END_REGION

REGION Network 2: EM - Resetting State Complete
   RUNG wire#powerrail
      Contact( "EM02".PackML_Sts.Alarm.sts_Resetting_SC )
      wire#w1
      Contact( "EM02".PackML_Sts.CM01.sts_Resetting_SC )
      wire#w2
      Contact( "EM02".PackML_Sts.CM02.sts_Resetting_SC )
      wire#w3
      Contact( "EM02".PackML_Sts.CM03.sts_Resetting_SC )
      wire#w4
      Contact( "EM02".PackML_Sts.CM04.sts_Resetting_SC )
      wire#w5
      Contact( "EM02".PackML_Sts.CM05.sts_Resetting_SC )
      wire#w6
      Contact( "EM02".PackML_Sts.CM06.sts_Resetting_SC )
      wire#w7
      Contact( "EM02".PackML_Sts.CM07.sts_Resetting_SC )
      wire#w8
      Contact( "EM02".PackML_Sts.CM08.sts_Resetting_SC )
      wire#w9
      Contact( "EM02".PackML_Sts.CM09.sts_Resetting_SC )
      wire#w10
      Contact( "EM02".PackML_Sts.CM10.sts_Resetting_SC )
      wire#w11
      Coil( "EM02".PackML_Sts.Unit.sts_Resetting_SC )
   END_RUNG
   RUNG wire#powerrail
      I_Contact( "EM02".PackML_Sts.Alarm.moduleActive )
   END_RUNG wire#w1
   RUNG wire#w1
      I_Contact( "EM02".PackML_Sts.CM01.moduleActive )
   END_RUNG wire#w2
   RUNG wire#w2
      I_Contact( "EM02".PackML_Sts.CM02.moduleActive )
   END_RUNG wire#w3
   RUNG wire#w3
      I_Contact( "EM02".PackML_Sts.CM03.moduleActive )
   END_RUNG wire#w4
   RUNG wire#w4
      I_Contact( "EM02".PackML_Sts.CM04.moduleActive )
   END_RUNG wire#w5
   RUNG wire#w5
      I_Contact( "EM02".PackML_Sts.CM05.moduleActive )
   END_RUNG wire#w6
   RUNG wire#w6
      I_Contact( "EM02".PackML_Sts.CM06.moduleActive )
   END_RUNG wire#w7
   RUNG wire#w7
      I_Contact( "EM02".PackML_Sts.CM07.moduleActive )
   END_RUNG wire#w8
   RUNG wire#w8
      I_Contact( "EM02".PackML_Sts.CM08.moduleActive )
   END_RUNG wire#w9
   RUNG wire#w9
      I_Contact( "EM02".PackML_Sts.CM09.moduleActive )
   END_RUNG wire#w10
   RUNG wire#w10
      I_Contact( "EM02".PackML_Sts.CM10.moduleActive )
   END_RUNG wire#w11
   // the same network as SCL:
   "EM02".PackML_Sts.Unit.sts_Resetting_SC := ("EM02".PackML_Sts.Alarm.sts_Resetting_SC OR NOT "EM02".PackML_Sts.Alarm.moduleActive) AND ("EM02".PackML_Sts.CM01.sts_Resetting_SC OR NOT "EM02".PackML_Sts.CM01.moduleActive) AND ("EM02".PackML_Sts.CM02.sts_Resetting_SC OR NOT "EM02".PackML_Sts.CM02.moduleActive) AND ("EM02".PackML_Sts.CM03.sts_Resetting_SC OR NOT "EM02".PackML_Sts.CM03.moduleActive) AND ("EM02".PackML_Sts.CM04.sts_Resetting_SC OR NOT "EM02".PackML_Sts.CM04.moduleActive) AND ("EM02".PackML_Sts.CM05.sts_Resetting_SC OR NOT "EM02".PackML_Sts.CM05.moduleActive) AND ("EM02".PackML_Sts.CM06.sts_Resetting_SC OR NOT "EM02".PackML_Sts.CM06.moduleActive) AND ("EM02".PackML_Sts.CM07.sts_Resetting_SC OR NOT "EM02".PackML_Sts.CM07.moduleActive) AND ("EM02".PackML_Sts.CM08.sts_Resetting_SC OR NOT "EM02".PackML_Sts.CM08.moduleActive) AND ("EM02".PackML_Sts.CM09.sts_Resetting_SC OR NOT "EM02".PackML_Sts.CM09.moduleActive) AND ("EM02".PackML_Sts.CM10.sts_Resetting_SC OR NOT "EM02".PackML_Sts.CM10.moduleActive);
END_REGION

REGION Network 3: EM - Start Command
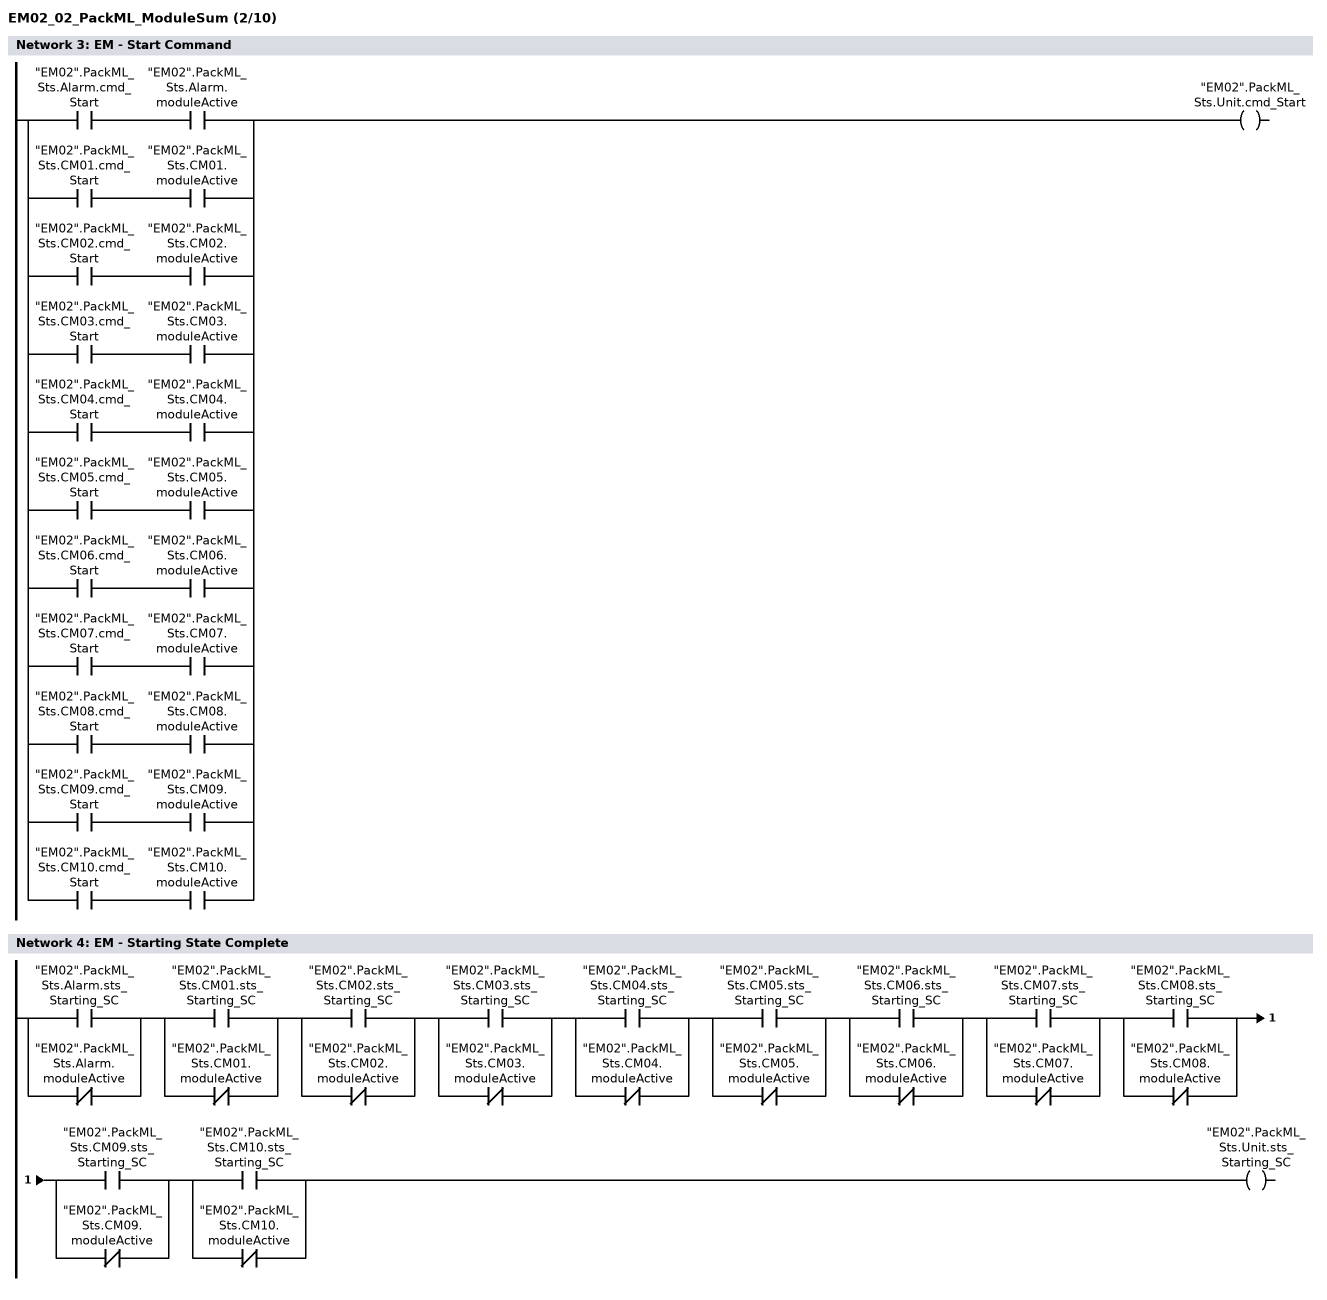
   RUNG wire#powerrail
      Contact( "EM02".PackML_Sts.Alarm.cmd_Start )
      Contact( "EM02".PackML_Sts.Alarm.moduleActive )
      wire#w1
      Coil( "EM02".PackML_Sts.Unit.cmd_Start )
   END_RUNG
   RUNG wire#powerrail
      Contact( "EM02".PackML_Sts.CM01.cmd_Start )
      Contact( "EM02".PackML_Sts.CM01.moduleActive )
   END_RUNG wire#w1
   RUNG wire#powerrail
      Contact( "EM02".PackML_Sts.CM02.cmd_Start )
      Contact( "EM02".PackML_Sts.CM02.moduleActive )
   END_RUNG wire#w1
   RUNG wire#powerrail
      Contact( "EM02".PackML_Sts.CM03.cmd_Start )
      Contact( "EM02".PackML_Sts.CM03.moduleActive )
   END_RUNG wire#w1
   RUNG wire#powerrail
      Contact( "EM02".PackML_Sts.CM04.cmd_Start )
      Contact( "EM02".PackML_Sts.CM04.moduleActive )
   END_RUNG wire#w1
   RUNG wire#powerrail
      Contact( "EM02".PackML_Sts.CM05.cmd_Start )
      Contact( "EM02".PackML_Sts.CM05.moduleActive )
   END_RUNG wire#w1
   RUNG wire#powerrail
      Contact( "EM02".PackML_Sts.CM06.cmd_Start )
      Contact( "EM02".PackML_Sts.CM06.moduleActive )
   END_RUNG wire#w1
   RUNG wire#powerrail
      Contact( "EM02".PackML_Sts.CM07.cmd_Start )
      Contact( "EM02".PackML_Sts.CM07.moduleActive )
   END_RUNG wire#w1
   RUNG wire#powerrail
      Contact( "EM02".PackML_Sts.CM08.cmd_Start )
      Contact( "EM02".PackML_Sts.CM08.moduleActive )
   END_RUNG wire#w1
   RUNG wire#powerrail
      Contact( "EM02".PackML_Sts.CM09.cmd_Start )
      Contact( "EM02".PackML_Sts.CM09.moduleActive )
   END_RUNG wire#w1
   RUNG wire#powerrail
      Contact( "EM02".PackML_Sts.CM10.cmd_Start )
      Contact( "EM02".PackML_Sts.CM10.moduleActive )
   END_RUNG wire#w1
   // the same network as SCL:
   "EM02".PackML_Sts.Unit.cmd_Start := ("EM02".PackML_Sts.Alarm.cmd_Start AND "EM02".PackML_Sts.Alarm.moduleActive) OR ("EM02".PackML_Sts.CM01.cmd_Start AND "EM02".PackML_Sts.CM01.moduleActive) OR ("EM02".PackML_Sts.CM02.cmd_Start AND "EM02".PackML_Sts.CM02.moduleActive) OR ("EM02".PackML_Sts.CM03.cmd_Start AND "EM02".PackML_Sts.CM03.moduleActive) OR ("EM02".PackML_Sts.CM04.cmd_Start AND "EM02".PackML_Sts.CM04.moduleActive) OR ("EM02".PackML_Sts.CM05.cmd_Start AND "EM02".PackML_Sts.CM05.moduleActive) OR ("EM02".PackML_Sts.CM06.cmd_Start AND "EM02".PackML_Sts.CM06.moduleActive) OR ("EM02".PackML_Sts.CM07.cmd_Start AND "EM02".PackML_Sts.CM07.moduleActive) OR ("EM02".PackML_Sts.CM08.cmd_Start AND "EM02".PackML_Sts.CM08.moduleActive) OR ("EM02".PackML_Sts.CM09.cmd_Start AND "EM02".PackML_Sts.CM09.moduleActive) OR ("EM02".PackML_Sts.CM10.cmd_Start AND "EM02".PackML_Sts.CM10.moduleActive);
END_REGION

REGION Network 4: EM - Starting State Complete
   RUNG wire#powerrail
      Contact( "EM02".PackML_Sts.Alarm.sts_Starting_SC )
      wire#w1
      Contact( "EM02".PackML_Sts.CM01.sts_Starting_SC )
      wire#w2
      Contact( "EM02".PackML_Sts.CM02.sts_Starting_SC )
      wire#w3
      Contact( "EM02".PackML_Sts.CM03.sts_Starting_SC )
      wire#w4
      Contact( "EM02".PackML_Sts.CM04.sts_Starting_SC )
      wire#w5
      Contact( "EM02".PackML_Sts.CM05.sts_Starting_SC )
      wire#w6
      Contact( "EM02".PackML_Sts.CM06.sts_Starting_SC )
      wire#w7
      Contact( "EM02".PackML_Sts.CM07.sts_Starting_SC )
      wire#w8
      Contact( "EM02".PackML_Sts.CM08.sts_Starting_SC )
      wire#w9
      Contact( "EM02".PackML_Sts.CM09.sts_Starting_SC )
      wire#w10
      Contact( "EM02".PackML_Sts.CM10.sts_Starting_SC )
      wire#w11
      Coil( "EM02".PackML_Sts.Unit.sts_Starting_SC )
   END_RUNG
   RUNG wire#powerrail
      I_Contact( "EM02".PackML_Sts.Alarm.moduleActive )
   END_RUNG wire#w1
   RUNG wire#w1
      I_Contact( "EM02".PackML_Sts.CM01.moduleActive )
   END_RUNG wire#w2
   RUNG wire#w2
      I_Contact( "EM02".PackML_Sts.CM02.moduleActive )
   END_RUNG wire#w3
   RUNG wire#w3
      I_Contact( "EM02".PackML_Sts.CM03.moduleActive )
   END_RUNG wire#w4
   RUNG wire#w4
      I_Contact( "EM02".PackML_Sts.CM04.moduleActive )
   END_RUNG wire#w5
   RUNG wire#w5
      I_Contact( "EM02".PackML_Sts.CM05.moduleActive )
   END_RUNG wire#w6
   RUNG wire#w6
      I_Contact( "EM02".PackML_Sts.CM06.moduleActive )
   END_RUNG wire#w7
   RUNG wire#w7
      I_Contact( "EM02".PackML_Sts.CM07.moduleActive )
   END_RUNG wire#w8
   RUNG wire#w8
      I_Contact( "EM02".PackML_Sts.CM08.moduleActive )
   END_RUNG wire#w9
   RUNG wire#w9
      I_Contact( "EM02".PackML_Sts.CM09.moduleActive )
   END_RUNG wire#w10
   RUNG wire#w10
      I_Contact( "EM02".PackML_Sts.CM10.moduleActive )
   END_RUNG wire#w11
   // the same network as SCL:
   "EM02".PackML_Sts.Unit.sts_Starting_SC := ("EM02".PackML_Sts.Alarm.sts_Starting_SC OR NOT "EM02".PackML_Sts.Alarm.moduleActive) AND ("EM02".PackML_Sts.CM01.sts_Starting_SC OR NOT "EM02".PackML_Sts.CM01.moduleActive) AND ("EM02".PackML_Sts.CM02.sts_Starting_SC OR NOT "EM02".PackML_Sts.CM02.moduleActive) AND ("EM02".PackML_Sts.CM03.sts_Starting_SC OR NOT "EM02".PackML_Sts.CM03.moduleActive) AND ("EM02".PackML_Sts.CM04.sts_Starting_SC OR NOT "EM02".PackML_Sts.CM04.moduleActive) AND ("EM02".PackML_Sts.CM05.sts_Starting_SC OR NOT "EM02".PackML_Sts.CM05.moduleActive) AND ("EM02".PackML_Sts.CM06.sts_Starting_SC OR NOT "EM02".PackML_Sts.CM06.moduleActive) AND ("EM02".PackML_Sts.CM07.sts_Starting_SC OR NOT "EM02".PackML_Sts.CM07.moduleActive) AND ("EM02".PackML_Sts.CM08.sts_Starting_SC OR NOT "EM02".PackML_Sts.CM08.moduleActive) AND ("EM02".PackML_Sts.CM09.sts_Starting_SC OR NOT "EM02".PackML_Sts.CM09.moduleActive) AND ("EM02".PackML_Sts.CM10.sts_Starting_SC OR NOT "EM02".PackML_Sts.CM10.moduleActive);
END_REGION

REGION Network 5: EM - Stop Command
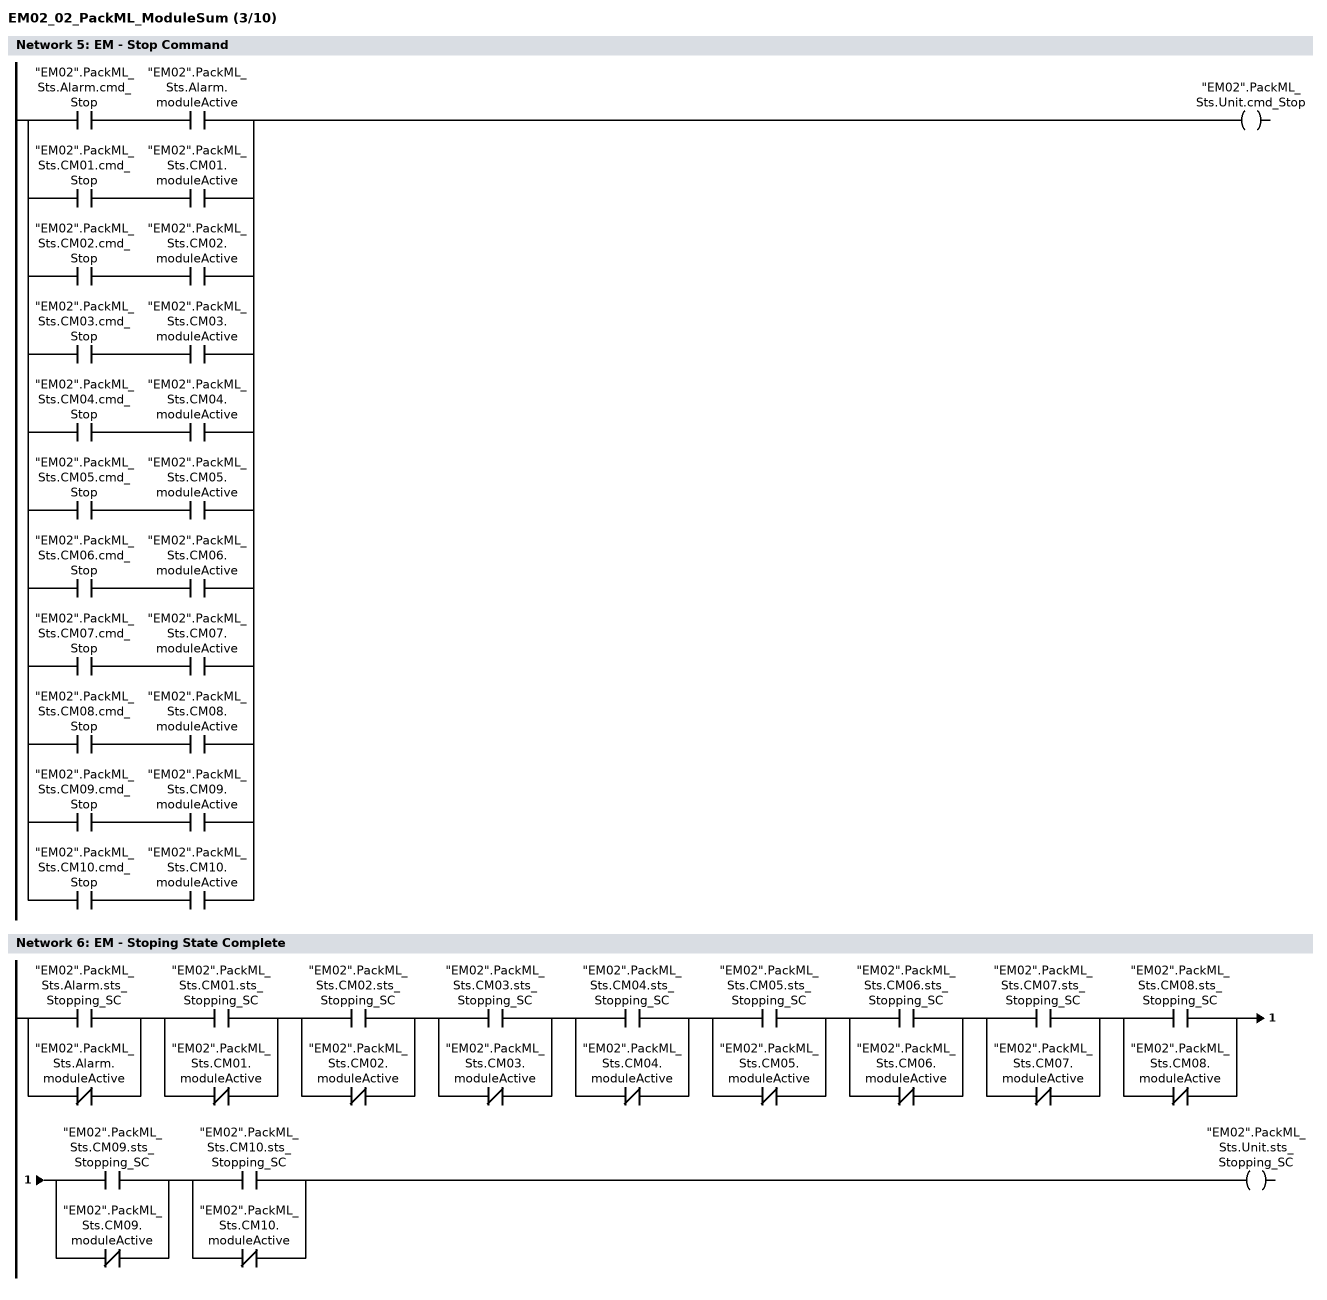
   RUNG wire#powerrail
      Contact( "EM02".PackML_Sts.Alarm.cmd_Stop )
      Contact( "EM02".PackML_Sts.Alarm.moduleActive )
      wire#w1
      Coil( "EM02".PackML_Sts.Unit.cmd_Stop )
   END_RUNG
   RUNG wire#powerrail
      Contact( "EM02".PackML_Sts.CM01.cmd_Stop )
      Contact( "EM02".PackML_Sts.CM01.moduleActive )
   END_RUNG wire#w1
   RUNG wire#powerrail
      Contact( "EM02".PackML_Sts.CM02.cmd_Stop )
      Contact( "EM02".PackML_Sts.CM02.moduleActive )
   END_RUNG wire#w1
   RUNG wire#powerrail
      Contact( "EM02".PackML_Sts.CM03.cmd_Stop )
      Contact( "EM02".PackML_Sts.CM03.moduleActive )
   END_RUNG wire#w1
   RUNG wire#powerrail
      Contact( "EM02".PackML_Sts.CM04.cmd_Stop )
      Contact( "EM02".PackML_Sts.CM04.moduleActive )
   END_RUNG wire#w1
   RUNG wire#powerrail
      Contact( "EM02".PackML_Sts.CM05.cmd_Stop )
      Contact( "EM02".PackML_Sts.CM05.moduleActive )
   END_RUNG wire#w1
   RUNG wire#powerrail
      Contact( "EM02".PackML_Sts.CM06.cmd_Stop )
      Contact( "EM02".PackML_Sts.CM06.moduleActive )
   END_RUNG wire#w1
   RUNG wire#powerrail
      Contact( "EM02".PackML_Sts.CM07.cmd_Stop )
      Contact( "EM02".PackML_Sts.CM07.moduleActive )
   END_RUNG wire#w1
   RUNG wire#powerrail
      Contact( "EM02".PackML_Sts.CM08.cmd_Stop )
      Contact( "EM02".PackML_Sts.CM08.moduleActive )
   END_RUNG wire#w1
   RUNG wire#powerrail
      Contact( "EM02".PackML_Sts.CM09.cmd_Stop )
      Contact( "EM02".PackML_Sts.CM09.moduleActive )
   END_RUNG wire#w1
   RUNG wire#powerrail
      Contact( "EM02".PackML_Sts.CM10.cmd_Stop )
      Contact( "EM02".PackML_Sts.CM10.moduleActive )
   END_RUNG wire#w1
   // the same network as SCL:
   "EM02".PackML_Sts.Unit.cmd_Stop := ("EM02".PackML_Sts.Alarm.cmd_Stop AND "EM02".PackML_Sts.Alarm.moduleActive) OR ("EM02".PackML_Sts.CM01.cmd_Stop AND "EM02".PackML_Sts.CM01.moduleActive) OR ("EM02".PackML_Sts.CM02.cmd_Stop AND "EM02".PackML_Sts.CM02.moduleActive) OR ("EM02".PackML_Sts.CM03.cmd_Stop AND "EM02".PackML_Sts.CM03.moduleActive) OR ("EM02".PackML_Sts.CM04.cmd_Stop AND "EM02".PackML_Sts.CM04.moduleActive) OR ("EM02".PackML_Sts.CM05.cmd_Stop AND "EM02".PackML_Sts.CM05.moduleActive) OR ("EM02".PackML_Sts.CM06.cmd_Stop AND "EM02".PackML_Sts.CM06.moduleActive) OR ("EM02".PackML_Sts.CM07.cmd_Stop AND "EM02".PackML_Sts.CM07.moduleActive) OR ("EM02".PackML_Sts.CM08.cmd_Stop AND "EM02".PackML_Sts.CM08.moduleActive) OR ("EM02".PackML_Sts.CM09.cmd_Stop AND "EM02".PackML_Sts.CM09.moduleActive) OR ("EM02".PackML_Sts.CM10.cmd_Stop AND "EM02".PackML_Sts.CM10.moduleActive);
END_REGION

REGION Network 6: EM - Stoping State Complete
   RUNG wire#powerrail
      Contact( "EM02".PackML_Sts.Alarm.sts_Stopping_SC )
      wire#w1
      Contact( "EM02".PackML_Sts.CM01.sts_Stopping_SC )
      wire#w2
      Contact( "EM02".PackML_Sts.CM02.sts_Stopping_SC )
      wire#w3
      Contact( "EM02".PackML_Sts.CM03.sts_Stopping_SC )
      wire#w4
      Contact( "EM02".PackML_Sts.CM04.sts_Stopping_SC )
      wire#w5
      Contact( "EM02".PackML_Sts.CM05.sts_Stopping_SC )
      wire#w6
      Contact( "EM02".PackML_Sts.CM06.sts_Stopping_SC )
      wire#w7
      Contact( "EM02".PackML_Sts.CM07.sts_Stopping_SC )
      wire#w8
      Contact( "EM02".PackML_Sts.CM08.sts_Stopping_SC )
      wire#w9
      Contact( "EM02".PackML_Sts.CM09.sts_Stopping_SC )
      wire#w10
      Contact( "EM02".PackML_Sts.CM10.sts_Stopping_SC )
      wire#w11
      Coil( "EM02".PackML_Sts.Unit.sts_Stopping_SC )
   END_RUNG
   RUNG wire#powerrail
      I_Contact( "EM02".PackML_Sts.Alarm.moduleActive )
   END_RUNG wire#w1
   RUNG wire#w1
      I_Contact( "EM02".PackML_Sts.CM01.moduleActive )
   END_RUNG wire#w2
   RUNG wire#w2
      I_Contact( "EM02".PackML_Sts.CM02.moduleActive )
   END_RUNG wire#w3
   RUNG wire#w3
      I_Contact( "EM02".PackML_Sts.CM03.moduleActive )
   END_RUNG wire#w4
   RUNG wire#w4
      I_Contact( "EM02".PackML_Sts.CM04.moduleActive )
   END_RUNG wire#w5
   RUNG wire#w5
      I_Contact( "EM02".PackML_Sts.CM05.moduleActive )
   END_RUNG wire#w6
   RUNG wire#w6
      I_Contact( "EM02".PackML_Sts.CM06.moduleActive )
   END_RUNG wire#w7
   RUNG wire#w7
      I_Contact( "EM02".PackML_Sts.CM07.moduleActive )
   END_RUNG wire#w8
   RUNG wire#w8
      I_Contact( "EM02".PackML_Sts.CM08.moduleActive )
   END_RUNG wire#w9
   RUNG wire#w9
      I_Contact( "EM02".PackML_Sts.CM09.moduleActive )
   END_RUNG wire#w10
   RUNG wire#w10
      I_Contact( "EM02".PackML_Sts.CM10.moduleActive )
   END_RUNG wire#w11
   // the same network as SCL:
   "EM02".PackML_Sts.Unit.sts_Stopping_SC := ("EM02".PackML_Sts.Alarm.sts_Stopping_SC OR NOT "EM02".PackML_Sts.Alarm.moduleActive) AND ("EM02".PackML_Sts.CM01.sts_Stopping_SC OR NOT "EM02".PackML_Sts.CM01.moduleActive) AND ("EM02".PackML_Sts.CM02.sts_Stopping_SC OR NOT "EM02".PackML_Sts.CM02.moduleActive) AND ("EM02".PackML_Sts.CM03.sts_Stopping_SC OR NOT "EM02".PackML_Sts.CM03.moduleActive) AND ("EM02".PackML_Sts.CM04.sts_Stopping_SC OR NOT "EM02".PackML_Sts.CM04.moduleActive) AND ("EM02".PackML_Sts.CM05.sts_Stopping_SC OR NOT "EM02".PackML_Sts.CM05.moduleActive) AND ("EM02".PackML_Sts.CM06.sts_Stopping_SC OR NOT "EM02".PackML_Sts.CM06.moduleActive) AND ("EM02".PackML_Sts.CM07.sts_Stopping_SC OR NOT "EM02".PackML_Sts.CM07.moduleActive) AND ("EM02".PackML_Sts.CM08.sts_Stopping_SC OR NOT "EM02".PackML_Sts.CM08.moduleActive) AND ("EM02".PackML_Sts.CM09.sts_Stopping_SC OR NOT "EM02".PackML_Sts.CM09.moduleActive) AND ("EM02".PackML_Sts.CM10.sts_Stopping_SC OR NOT "EM02".PackML_Sts.CM10.moduleActive);
END_REGION

REGION Network 7: EM - Hold Command
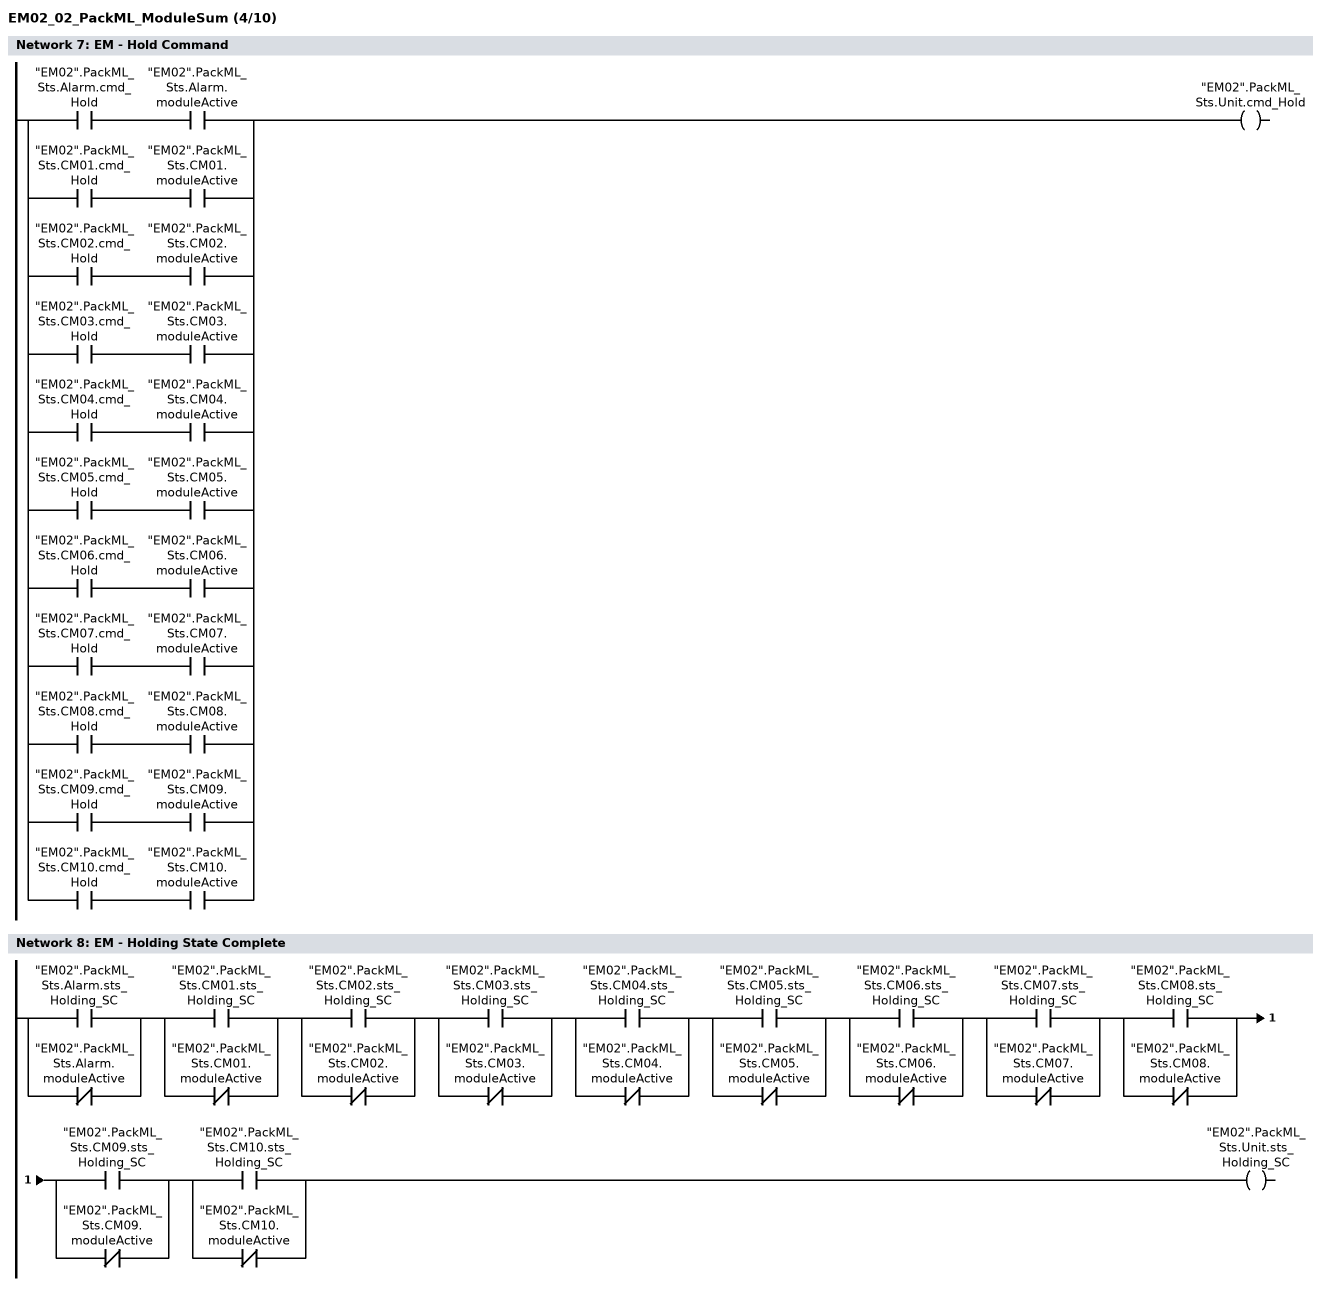
   RUNG wire#powerrail
      Contact( "EM02".PackML_Sts.Alarm.cmd_Hold )
      Contact( "EM02".PackML_Sts.Alarm.moduleActive )
      wire#w1
      Coil( "EM02".PackML_Sts.Unit.cmd_Hold )
   END_RUNG
   RUNG wire#powerrail
      Contact( "EM02".PackML_Sts.CM01.cmd_Hold )
      Contact( "EM02".PackML_Sts.CM01.moduleActive )
   END_RUNG wire#w1
   RUNG wire#powerrail
      Contact( "EM02".PackML_Sts.CM02.cmd_Hold )
      Contact( "EM02".PackML_Sts.CM02.moduleActive )
   END_RUNG wire#w1
   RUNG wire#powerrail
      Contact( "EM02".PackML_Sts.CM03.cmd_Hold )
      Contact( "EM02".PackML_Sts.CM03.moduleActive )
   END_RUNG wire#w1
   RUNG wire#powerrail
      Contact( "EM02".PackML_Sts.CM04.cmd_Hold )
      Contact( "EM02".PackML_Sts.CM04.moduleActive )
   END_RUNG wire#w1
   RUNG wire#powerrail
      Contact( "EM02".PackML_Sts.CM05.cmd_Hold )
      Contact( "EM02".PackML_Sts.CM05.moduleActive )
   END_RUNG wire#w1
   RUNG wire#powerrail
      Contact( "EM02".PackML_Sts.CM06.cmd_Hold )
      Contact( "EM02".PackML_Sts.CM06.moduleActive )
   END_RUNG wire#w1
   RUNG wire#powerrail
      Contact( "EM02".PackML_Sts.CM07.cmd_Hold )
      Contact( "EM02".PackML_Sts.CM07.moduleActive )
   END_RUNG wire#w1
   RUNG wire#powerrail
      Contact( "EM02".PackML_Sts.CM08.cmd_Hold )
      Contact( "EM02".PackML_Sts.CM08.moduleActive )
   END_RUNG wire#w1
   RUNG wire#powerrail
      Contact( "EM02".PackML_Sts.CM09.cmd_Hold )
      Contact( "EM02".PackML_Sts.CM09.moduleActive )
   END_RUNG wire#w1
   RUNG wire#powerrail
      Contact( "EM02".PackML_Sts.CM10.cmd_Hold )
      Contact( "EM02".PackML_Sts.CM10.moduleActive )
   END_RUNG wire#w1
   // the same network as SCL:
   "EM02".PackML_Sts.Unit.cmd_Hold := ("EM02".PackML_Sts.Alarm.cmd_Hold AND "EM02".PackML_Sts.Alarm.moduleActive) OR ("EM02".PackML_Sts.CM01.cmd_Hold AND "EM02".PackML_Sts.CM01.moduleActive) OR ("EM02".PackML_Sts.CM02.cmd_Hold AND "EM02".PackML_Sts.CM02.moduleActive) OR ("EM02".PackML_Sts.CM03.cmd_Hold AND "EM02".PackML_Sts.CM03.moduleActive) OR ("EM02".PackML_Sts.CM04.cmd_Hold AND "EM02".PackML_Sts.CM04.moduleActive) OR ("EM02".PackML_Sts.CM05.cmd_Hold AND "EM02".PackML_Sts.CM05.moduleActive) OR ("EM02".PackML_Sts.CM06.cmd_Hold AND "EM02".PackML_Sts.CM06.moduleActive) OR ("EM02".PackML_Sts.CM07.cmd_Hold AND "EM02".PackML_Sts.CM07.moduleActive) OR ("EM02".PackML_Sts.CM08.cmd_Hold AND "EM02".PackML_Sts.CM08.moduleActive) OR ("EM02".PackML_Sts.CM09.cmd_Hold AND "EM02".PackML_Sts.CM09.moduleActive) OR ("EM02".PackML_Sts.CM10.cmd_Hold AND "EM02".PackML_Sts.CM10.moduleActive);
END_REGION

REGION Network 8: EM - Holding State Complete
   RUNG wire#powerrail
      Contact( "EM02".PackML_Sts.Alarm.sts_Holding_SC )
      wire#w1
      Contact( "EM02".PackML_Sts.CM01.sts_Holding_SC )
      wire#w2
      Contact( "EM02".PackML_Sts.CM02.sts_Holding_SC )
      wire#w3
      Contact( "EM02".PackML_Sts.CM03.sts_Holding_SC )
      wire#w4
      Contact( "EM02".PackML_Sts.CM04.sts_Holding_SC )
      wire#w5
      Contact( "EM02".PackML_Sts.CM05.sts_Holding_SC )
      wire#w6
      Contact( "EM02".PackML_Sts.CM06.sts_Holding_SC )
      wire#w7
      Contact( "EM02".PackML_Sts.CM07.sts_Holding_SC )
      wire#w8
      Contact( "EM02".PackML_Sts.CM08.sts_Holding_SC )
      wire#w9
      Contact( "EM02".PackML_Sts.CM09.sts_Holding_SC )
      wire#w10
      Contact( "EM02".PackML_Sts.CM10.sts_Holding_SC )
      wire#w11
      Coil( "EM02".PackML_Sts.Unit.sts_Holding_SC )
   END_RUNG
   RUNG wire#powerrail
      I_Contact( "EM02".PackML_Sts.Alarm.moduleActive )
   END_RUNG wire#w1
   RUNG wire#w1
      I_Contact( "EM02".PackML_Sts.CM01.moduleActive )
   END_RUNG wire#w2
   RUNG wire#w2
      I_Contact( "EM02".PackML_Sts.CM02.moduleActive )
   END_RUNG wire#w3
   RUNG wire#w3
      I_Contact( "EM02".PackML_Sts.CM03.moduleActive )
   END_RUNG wire#w4
   RUNG wire#w4
      I_Contact( "EM02".PackML_Sts.CM04.moduleActive )
   END_RUNG wire#w5
   RUNG wire#w5
      I_Contact( "EM02".PackML_Sts.CM05.moduleActive )
   END_RUNG wire#w6
   RUNG wire#w6
      I_Contact( "EM02".PackML_Sts.CM06.moduleActive )
   END_RUNG wire#w7
   RUNG wire#w7
      I_Contact( "EM02".PackML_Sts.CM07.moduleActive )
   END_RUNG wire#w8
   RUNG wire#w8
      I_Contact( "EM02".PackML_Sts.CM08.moduleActive )
   END_RUNG wire#w9
   RUNG wire#w9
      I_Contact( "EM02".PackML_Sts.CM09.moduleActive )
   END_RUNG wire#w10
   RUNG wire#w10
      I_Contact( "EM02".PackML_Sts.CM10.moduleActive )
   END_RUNG wire#w11
   // the same network as SCL:
   "EM02".PackML_Sts.Unit.sts_Holding_SC := ("EM02".PackML_Sts.Alarm.sts_Holding_SC OR NOT "EM02".PackML_Sts.Alarm.moduleActive) AND ("EM02".PackML_Sts.CM01.sts_Holding_SC OR NOT "EM02".PackML_Sts.CM01.moduleActive) AND ("EM02".PackML_Sts.CM02.sts_Holding_SC OR NOT "EM02".PackML_Sts.CM02.moduleActive) AND ("EM02".PackML_Sts.CM03.sts_Holding_SC OR NOT "EM02".PackML_Sts.CM03.moduleActive) AND ("EM02".PackML_Sts.CM04.sts_Holding_SC OR NOT "EM02".PackML_Sts.CM04.moduleActive) AND ("EM02".PackML_Sts.CM05.sts_Holding_SC OR NOT "EM02".PackML_Sts.CM05.moduleActive) AND ("EM02".PackML_Sts.CM06.sts_Holding_SC OR NOT "EM02".PackML_Sts.CM06.moduleActive) AND ("EM02".PackML_Sts.CM07.sts_Holding_SC OR NOT "EM02".PackML_Sts.CM07.moduleActive) AND ("EM02".PackML_Sts.CM08.sts_Holding_SC OR NOT "EM02".PackML_Sts.CM08.moduleActive) AND ("EM02".PackML_Sts.CM09.sts_Holding_SC OR NOT "EM02".PackML_Sts.CM09.moduleActive) AND ("EM02".PackML_Sts.CM10.sts_Holding_SC OR NOT "EM02".PackML_Sts.CM10.moduleActive);
END_REGION

REGION Network 9: EM - UnHold Command
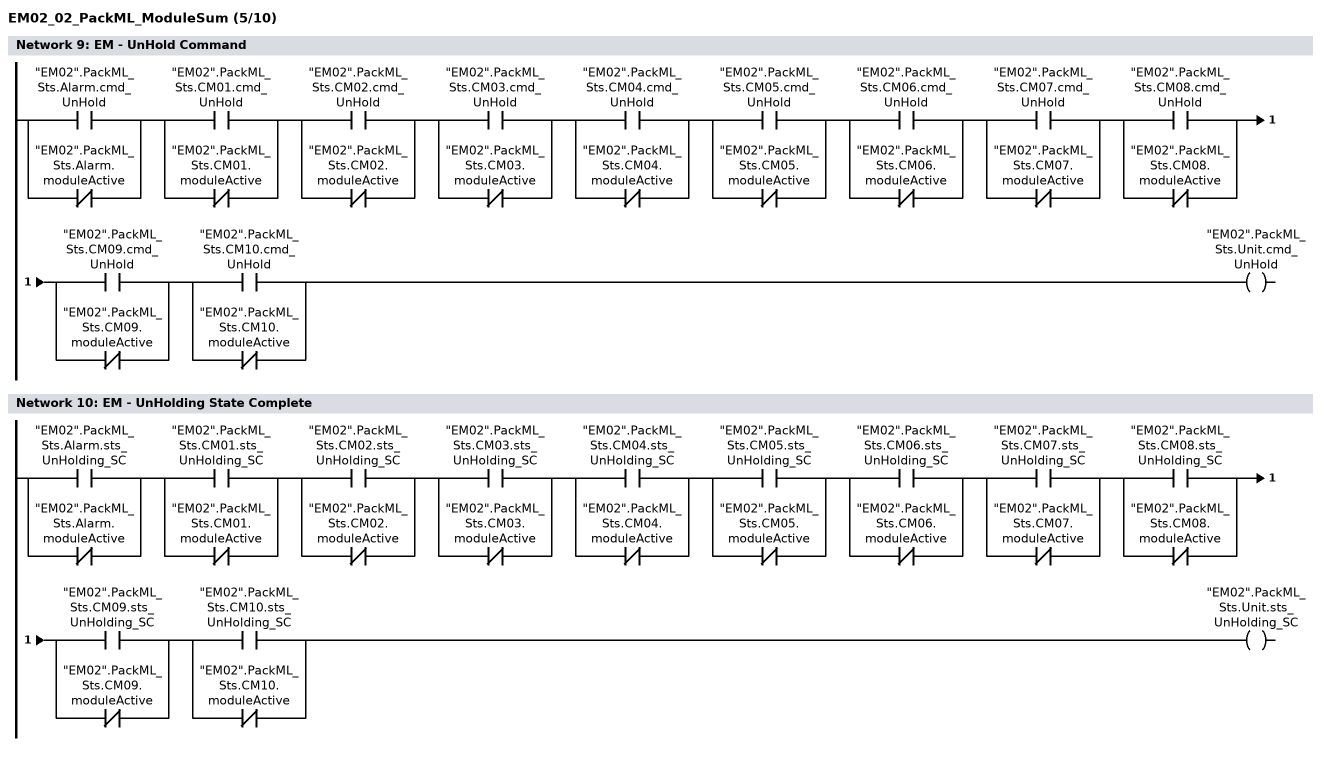
   RUNG wire#powerrail
      Contact( "EM02".PackML_Sts.Alarm.cmd_UnHold )
      wire#w1
      Contact( "EM02".PackML_Sts.CM01.cmd_UnHold )
      wire#w2
      Contact( "EM02".PackML_Sts.CM02.cmd_UnHold )
      wire#w3
      Contact( "EM02".PackML_Sts.CM03.cmd_UnHold )
      wire#w4
      Contact( "EM02".PackML_Sts.CM04.cmd_UnHold )
      wire#w5
      Contact( "EM02".PackML_Sts.CM05.cmd_UnHold )
      wire#w6
      Contact( "EM02".PackML_Sts.CM06.cmd_UnHold )
      wire#w7
      Contact( "EM02".PackML_Sts.CM07.cmd_UnHold )
      wire#w8
      Contact( "EM02".PackML_Sts.CM08.cmd_UnHold )
      wire#w9
      Contact( "EM02".PackML_Sts.CM09.cmd_UnHold )
      wire#w10
      Contact( "EM02".PackML_Sts.CM10.cmd_UnHold )
      wire#w11
      Coil( "EM02".PackML_Sts.Unit.cmd_UnHold )
   END_RUNG
   RUNG wire#powerrail
      I_Contact( "EM02".PackML_Sts.Alarm.moduleActive )
   END_RUNG wire#w1
   RUNG wire#w1
      I_Contact( "EM02".PackML_Sts.CM01.moduleActive )
   END_RUNG wire#w2
   RUNG wire#w2
      I_Contact( "EM02".PackML_Sts.CM02.moduleActive )
   END_RUNG wire#w3
   RUNG wire#w3
      I_Contact( "EM02".PackML_Sts.CM03.moduleActive )
   END_RUNG wire#w4
   RUNG wire#w4
      I_Contact( "EM02".PackML_Sts.CM04.moduleActive )
   END_RUNG wire#w5
   RUNG wire#w5
      I_Contact( "EM02".PackML_Sts.CM05.moduleActive )
   END_RUNG wire#w6
   RUNG wire#w6
      I_Contact( "EM02".PackML_Sts.CM06.moduleActive )
   END_RUNG wire#w7
   RUNG wire#w7
      I_Contact( "EM02".PackML_Sts.CM07.moduleActive )
   END_RUNG wire#w8
   RUNG wire#w8
      I_Contact( "EM02".PackML_Sts.CM08.moduleActive )
   END_RUNG wire#w9
   RUNG wire#w9
      I_Contact( "EM02".PackML_Sts.CM09.moduleActive )
   END_RUNG wire#w10
   RUNG wire#w10
      I_Contact( "EM02".PackML_Sts.CM10.moduleActive )
   END_RUNG wire#w11
   // the same network as SCL:
   "EM02".PackML_Sts.Unit.cmd_UnHold := ("EM02".PackML_Sts.Alarm.cmd_UnHold OR NOT "EM02".PackML_Sts.Alarm.moduleActive) AND ("EM02".PackML_Sts.CM01.cmd_UnHold OR NOT "EM02".PackML_Sts.CM01.moduleActive) AND ("EM02".PackML_Sts.CM02.cmd_UnHold OR NOT "EM02".PackML_Sts.CM02.moduleActive) AND ("EM02".PackML_Sts.CM03.cmd_UnHold OR NOT "EM02".PackML_Sts.CM03.moduleActive) AND ("EM02".PackML_Sts.CM04.cmd_UnHold OR NOT "EM02".PackML_Sts.CM04.moduleActive) AND ("EM02".PackML_Sts.CM05.cmd_UnHold OR NOT "EM02".PackML_Sts.CM05.moduleActive) AND ("EM02".PackML_Sts.CM06.cmd_UnHold OR NOT "EM02".PackML_Sts.CM06.moduleActive) AND ("EM02".PackML_Sts.CM07.cmd_UnHold OR NOT "EM02".PackML_Sts.CM07.moduleActive) AND ("EM02".PackML_Sts.CM08.cmd_UnHold OR NOT "EM02".PackML_Sts.CM08.moduleActive) AND ("EM02".PackML_Sts.CM09.cmd_UnHold OR NOT "EM02".PackML_Sts.CM09.moduleActive) AND ("EM02".PackML_Sts.CM10.cmd_UnHold OR NOT "EM02".PackML_Sts.CM10.moduleActive);
END_REGION
